(* Logix 5000 project; controller PLC_MCC1300_75F1 vendor 1 type 14 code 166 rev 32.11; software revision 32.04; part 17 of 83 *)
(* tags used below, declared in another part *)
   M302SpeedUp : MAC_SpeedUp;
   TMP_d : DINT;
   TMP_xPositioning : BOOL;
   TMP_xReverse : BOOL;
   TMP_xRun : BOOL;
   xAlwaysOFF : BOOL;
   Z300_Conveyor : UDT_StandConv[29];
   Z300_Conveyor_Conf : UDT_Conveyor_Config[29];
   Z300_Conveyor_HMW : MAC_Conveyor_ZC_HMW[29];
   Z300_Conveyor_IN_MOTION : MAC_Conveyor_ZC_IN_MOTION[29];
   Z301_HMR : MAC_Zone_ML_HMR;
(* CommandLogic, continued *)

ROUTINE M307BM1_Conveyor_Output   (* ladder *)
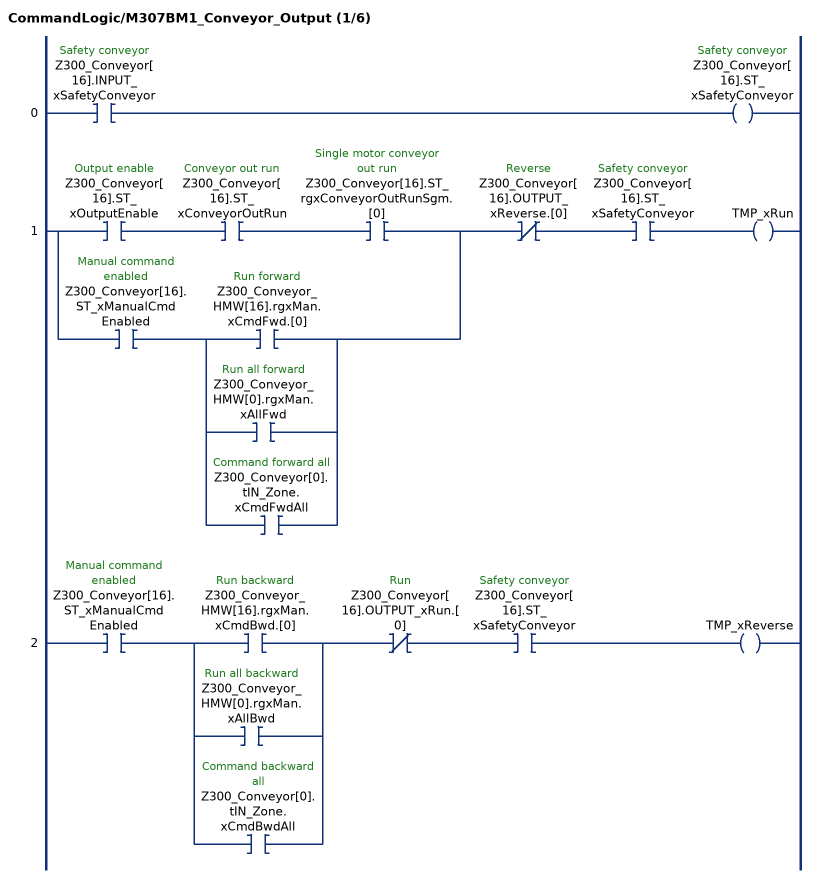
   0: XIC(Z300_Conveyor[16].INPUT_xSafetyConveyor)OTE(Z300_Conveyor[16].ST_xSafetyConveyor);
   1: [XIC(Z300_Conveyor[16].ST_xOutputEnable) XIC(Z300_Conveyor[16].ST_xConveyorOutRun) XIC(Z300_Conveyor[16].ST_rgxConveyorOutRunSgm.[0]) ,XIC(Z300_Conveyor[16].ST_xManualCmdEnabled) [XIC(Z300_Conveyor_HMW[16].rgxMan.xCmdFwd.[0]) ,XIC(Z300_Conveyor_HMW[0].rgxMan.xAllFwd) ,XIC(Z300_Conveyor[0].tIN_Zone.xCmdFwdAll) ] ]XIO(Z300_Conveyor[16].OUTPUT_xReverse.[0])XIC(Z300_Conveyor[16].ST_xSafetyConveyor)OTE(TMP_xRun);
   2: XIC(Z300_Conveyor[16].ST_xManualCmdEnabled)[XIC(Z300_Conveyor_HMW[16].rgxMan.xCmdBwd.[0]) ,XIC(Z300_Conveyor_HMW[0].rgxMan.xAllBwd) ,XIC(Z300_Conveyor[0].tIN_Zone.xCmdBwdAll) ]XIO(Z300_Conveyor[16].OUTPUT_xRun.[0])XIC(Z300_Conveyor[16].ST_xSafetyConveyor)OTE(TMP_xReverse);
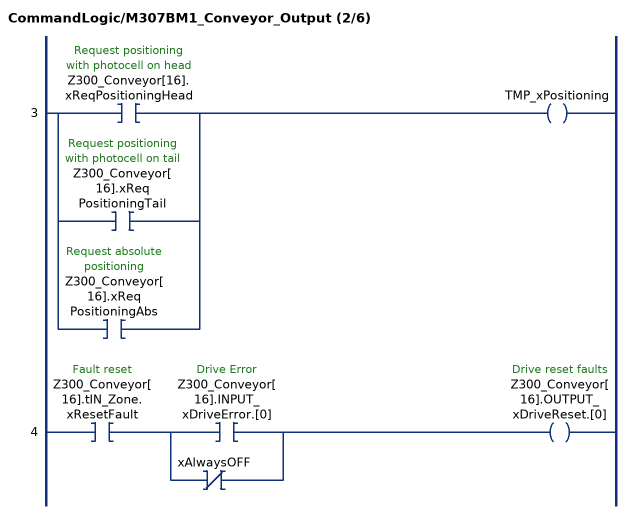
   3: [XIC(Z300_Conveyor[16].xReqPositioningHead) ,XIC(Z300_Conveyor[16].xReqPositioningTail) ,XIC(Z300_Conveyor[16].xReqPositioningAbs) ]OTE(TMP_xPositioning);
   4: XIC(Z300_Conveyor[16].tIN_Zone.xResetFault)[XIC(Z300_Conveyor[16].INPUT_xDriveError.[0]) ,XIO(xAlwaysOFF) ]OTE(Z300_Conveyor[16].OUTPUT_xDriveReset.[0]);
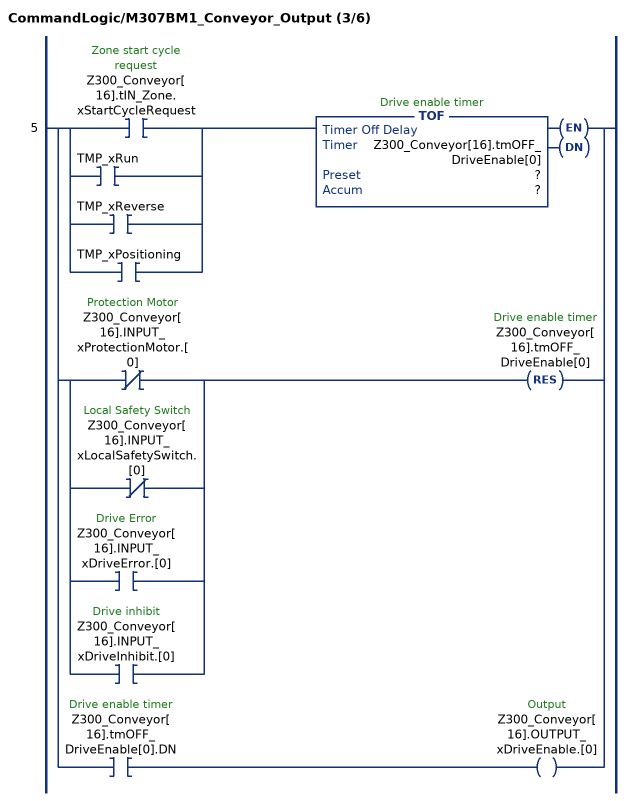
   5: [[XIC(Z300_Conveyor[16].tIN_Zone.xStartCycleRequest) ,XIC(TMP_xRun) ,XIC(TMP_xReverse) ,XIC(TMP_xPositioning) ] TOF(Z300_Conveyor[16].tmOFF_DriveEnable[0],?,?) ,[XIO(Z300_Conveyor[16].INPUT_xProtectionMotor.[0]) ,XIO(Z300_Conveyor[16].INPUT_xLocalSafetySwitch.[0]) ,XIC(Z300_Conveyor[16].INPUT_xDriveError.[0]) ,XIC(Z300_Conveyor[16].INPUT_xDriveInhibit.[0]) ] RES(Z300_Conveyor[16].tmOFF_DriveEnable[0]) ,XIC(Z300_Conveyor[16].tmOFF_DriveEnable[0].DN) OTE(Z300_Conveyor[16].OUTPUT_xDriveEnable.[0]) ];
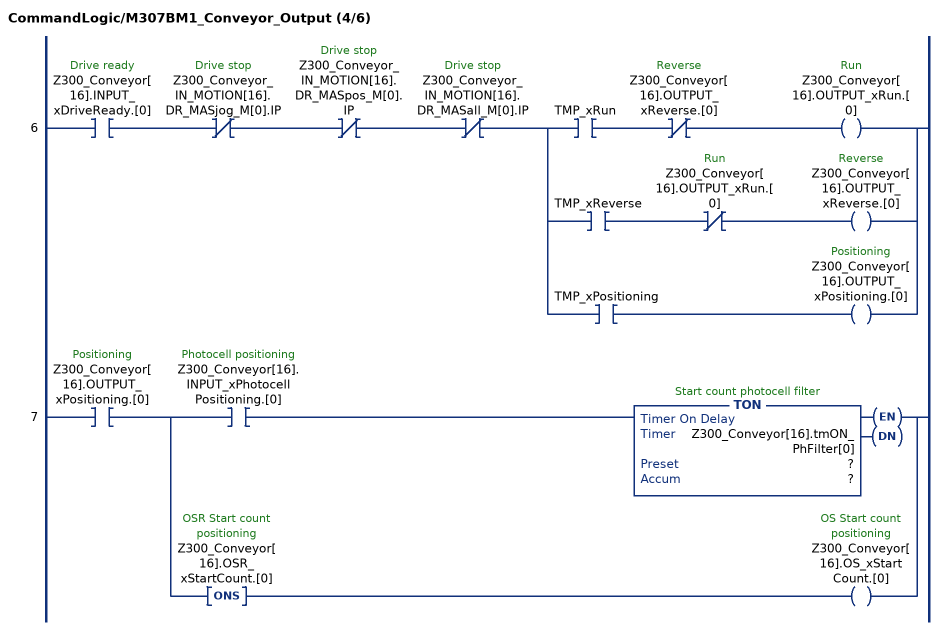
   6: XIC(Z300_Conveyor[16].INPUT_xDriveReady.[0])XIO(Z300_Conveyor_IN_MOTION[16].DR_MASjog_M[0].IP)XIO(Z300_Conveyor_IN_MOTION[16].DR_MASpos_M[0].IP)XIO(Z300_Conveyor_IN_MOTION[16].DR_MASall_M[0].IP)[XIC(TMP_xRun) XIO(Z300_Conveyor[16].OUTPUT_xReverse.[0]) OTE(Z300_Conveyor[16].OUTPUT_xRun.[0]) ,XIC(TMP_xReverse) XIO(Z300_Conveyor[16].OUTPUT_xRun.[0]) OTE(Z300_Conveyor[16].OUTPUT_xReverse.[0]) ,XIC(TMP_xPositioning) OTE(Z300_Conveyor[16].OUTPUT_xPositioning.[0]) ];
   7: XIC(Z300_Conveyor[16].OUTPUT_xPositioning.[0])[XIC(Z300_Conveyor[16].INPUT_xPhotocellPositioning.[0]) TON(Z300_Conveyor[16].tmON_PhFilter[0],?,?) ,ONS(Z300_Conveyor[16].OSR_xStartCount.[0]) OTE(Z300_Conveyor[16].OS_xStartCount.[0]) ];
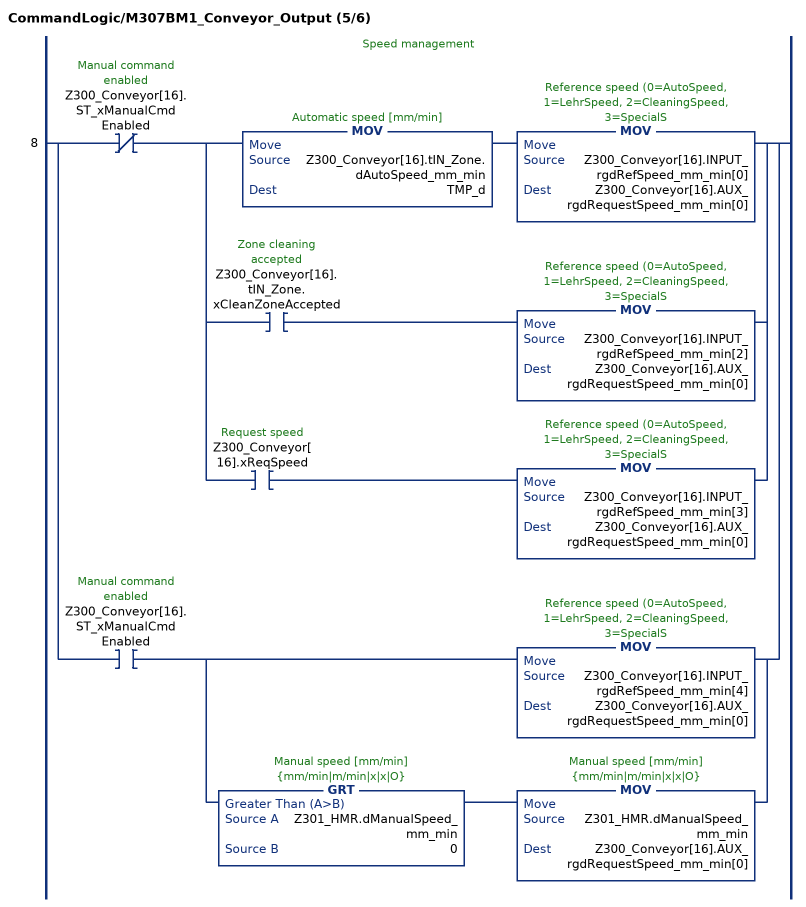
   // Speed management
   8: [XIO(Z300_Conveyor[16].ST_xManualCmdEnabled) [MOV(Z300_Conveyor[16].tIN_Zone.dAutoSpeed_mm_min,TMP_d) MOV(Z300_Conveyor[16].INPUT_rgdRefSpeed_mm_min[0],Z300_Conveyor[16].AUX_rgdRequestSpeed_mm_min[0]) ,XIC(Z300_Conveyor[16].tIN_Zone.xCleanZoneAccepted) MOV(Z300_Conveyor[16].INPUT_rgdRefSpeed_mm_min[2],Z300_Conveyor[16].AUX_rgdRequestSpeed_mm_min[0]) ,XIC(Z300_Conveyor[16].xReqSpeed) MOV(Z300_Conveyor[16].INPUT_rgdRefSpeed_mm_min[3],Z300_Conveyor[16].AUX_rgdRequestSpeed_mm_min[0]) ] ,XIC(Z300_Conveyor[16].ST_xManualCmdEnabled) [MOV(Z300_Conveyor[16].INPUT_rgdRefSpeed_mm_min[4],Z300_Conveyor[16].AUX_rgdRequestSpeed_mm_min[0]) ,GRT(Z301_HMR.dManualSpeed_mm_min,0) MOV(Z301_HMR.dManualSpeed_mm_min,Z300_Conveyor[16].AUX_rgdRequestSpeed_mm_min[0]) ] ];
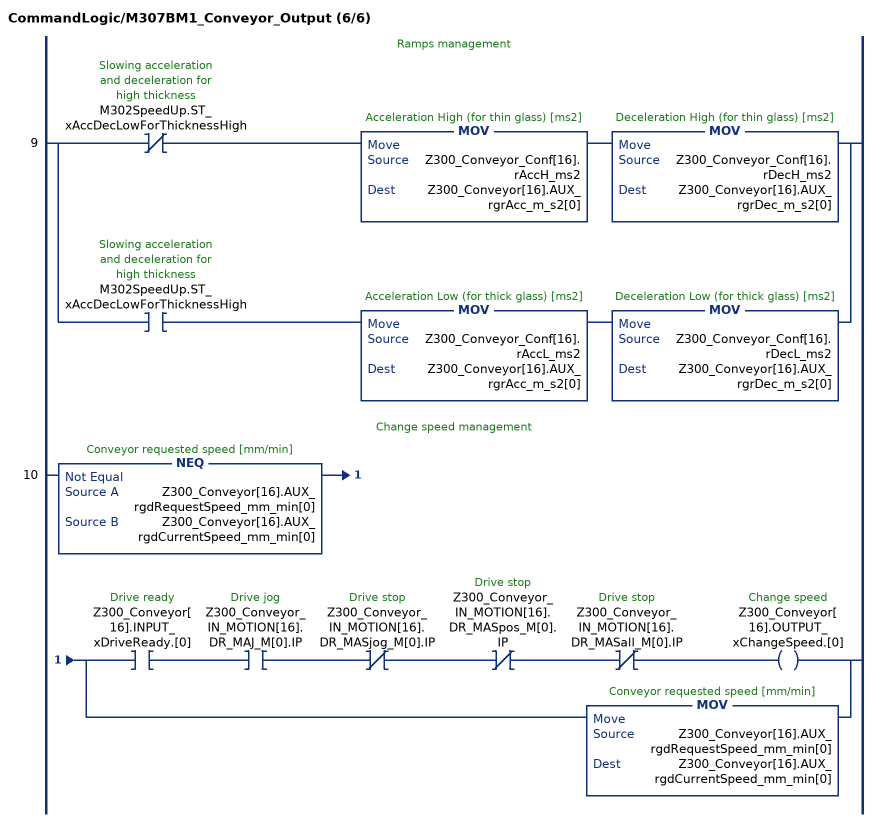
   // Ramps management
   9: [XIO(M302SpeedUp.ST_xAccDecLowForThicknessHigh) MOV(Z300_Conveyor_Conf[16].rAccH_ms2,Z300_Conveyor[16].AUX_rgrAcc_m_s2[0]) MOV(Z300_Conveyor_Conf[16].rDecH_ms2,Z300_Conveyor[16].AUX_rgrDec_m_s2[0]) ,XIC(M302SpeedUp.ST_xAccDecLowForThicknessHigh) MOV(Z300_Conveyor_Conf[16].rAccL_ms2,Z300_Conveyor[16].AUX_rgrAcc_m_s2[0]) MOV(Z300_Conveyor_Conf[16].rDecL_ms2,Z300_Conveyor[16].AUX_rgrDec_m_s2[0]) ];
   // Change speed management
   10: NEQ(Z300_Conveyor[16].AUX_rgdRequestSpeed_mm_min[0],Z300_Conveyor[16].AUX_rgdCurrentSpeed_mm_min[0])[XIC(Z300_Conveyor[16].INPUT_xDriveReady.[0]) XIC(Z300_Conveyor_IN_MOTION[16].DR_MAJ_M[0].IP) XIO(Z300_Conveyor_IN_MOTION[16].DR_MASjog_M[0].IP) XIO(Z300_Conveyor_IN_MOTION[16].DR_MASpos_M[0].IP) XIO(Z300_Conveyor_IN_MOTION[16].DR_MASall_M[0].IP) OTE(Z300_Conveyor[16].OUTPUT_xChangeSpeed.[0]) ,MOV(Z300_Conveyor[16].AUX_rgdRequestSpeed_mm_min[0],Z300_Conveyor[16].AUX_rgdCurrentSpeed_mm_min[0]) ];
END_ROUTINE

ROUTINE M307CM1_Conveyor_Output   (* ladder *)
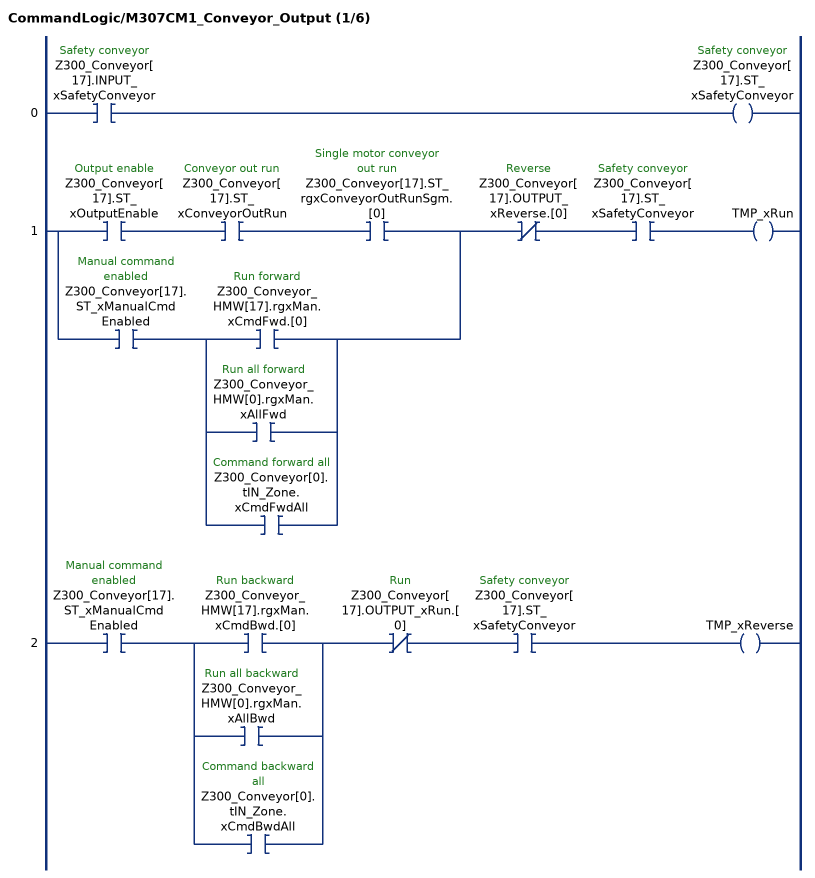
   0: XIC(Z300_Conveyor[17].INPUT_xSafetyConveyor)OTE(Z300_Conveyor[17].ST_xSafetyConveyor);
   1: [XIC(Z300_Conveyor[17].ST_xOutputEnable) XIC(Z300_Conveyor[17].ST_xConveyorOutRun) XIC(Z300_Conveyor[17].ST_rgxConveyorOutRunSgm.[0]) ,XIC(Z300_Conveyor[17].ST_xManualCmdEnabled) [XIC(Z300_Conveyor_HMW[17].rgxMan.xCmdFwd.[0]) ,XIC(Z300_Conveyor_HMW[0].rgxMan.xAllFwd) ,XIC(Z300_Conveyor[0].tIN_Zone.xCmdFwdAll) ] ]XIO(Z300_Conveyor[17].OUTPUT_xReverse.[0])XIC(Z300_Conveyor[17].ST_xSafetyConveyor)OTE(TMP_xRun);
   2: XIC(Z300_Conveyor[17].ST_xManualCmdEnabled)[XIC(Z300_Conveyor_HMW[17].rgxMan.xCmdBwd.[0]) ,XIC(Z300_Conveyor_HMW[0].rgxMan.xAllBwd) ,XIC(Z300_Conveyor[0].tIN_Zone.xCmdBwdAll) ]XIO(Z300_Conveyor[17].OUTPUT_xRun.[0])XIC(Z300_Conveyor[17].ST_xSafetyConveyor)OTE(TMP_xReverse);
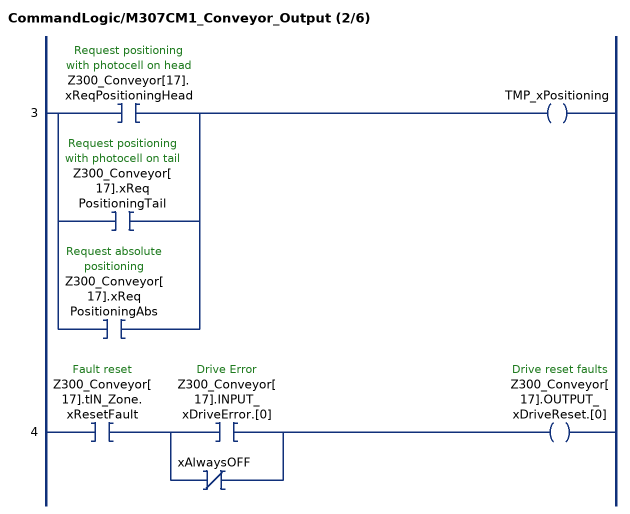
   3: [XIC(Z300_Conveyor[17].xReqPositioningHead) ,XIC(Z300_Conveyor[17].xReqPositioningTail) ,XIC(Z300_Conveyor[17].xReqPositioningAbs) ]OTE(TMP_xPositioning);
   4: XIC(Z300_Conveyor[17].tIN_Zone.xResetFault)[XIC(Z300_Conveyor[17].INPUT_xDriveError.[0]) ,XIO(xAlwaysOFF) ]OTE(Z300_Conveyor[17].OUTPUT_xDriveReset.[0]);
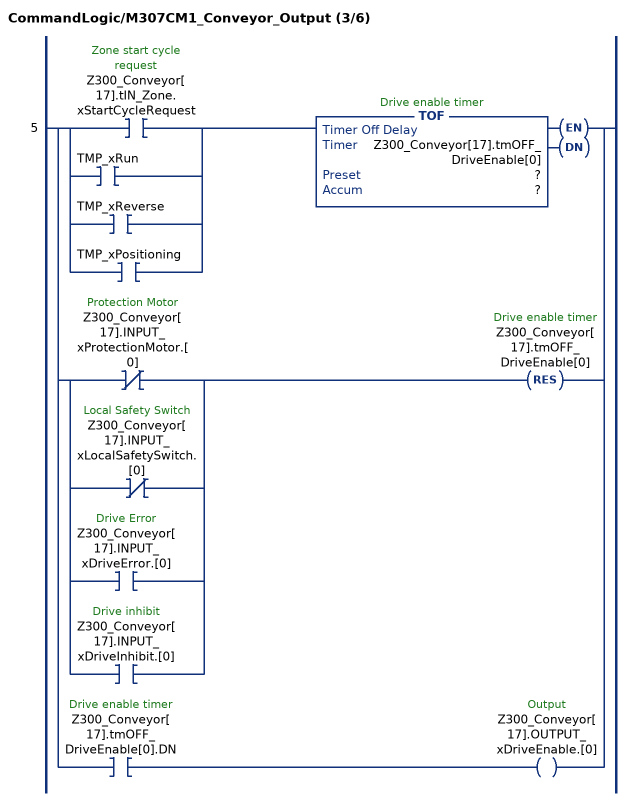
   5: [[XIC(Z300_Conveyor[17].tIN_Zone.xStartCycleRequest) ,XIC(TMP_xRun) ,XIC(TMP_xReverse) ,XIC(TMP_xPositioning) ] TOF(Z300_Conveyor[17].tmOFF_DriveEnable[0],?,?) ,[XIO(Z300_Conveyor[17].INPUT_xProtectionMotor.[0]) ,XIO(Z300_Conveyor[17].INPUT_xLocalSafetySwitch.[0]) ,XIC(Z300_Conveyor[17].INPUT_xDriveError.[0]) ,XIC(Z300_Conveyor[17].INPUT_xDriveInhibit.[0]) ] RES(Z300_Conveyor[17].tmOFF_DriveEnable[0]) ,XIC(Z300_Conveyor[17].tmOFF_DriveEnable[0].DN) OTE(Z300_Conveyor[17].OUTPUT_xDriveEnable.[0]) ];
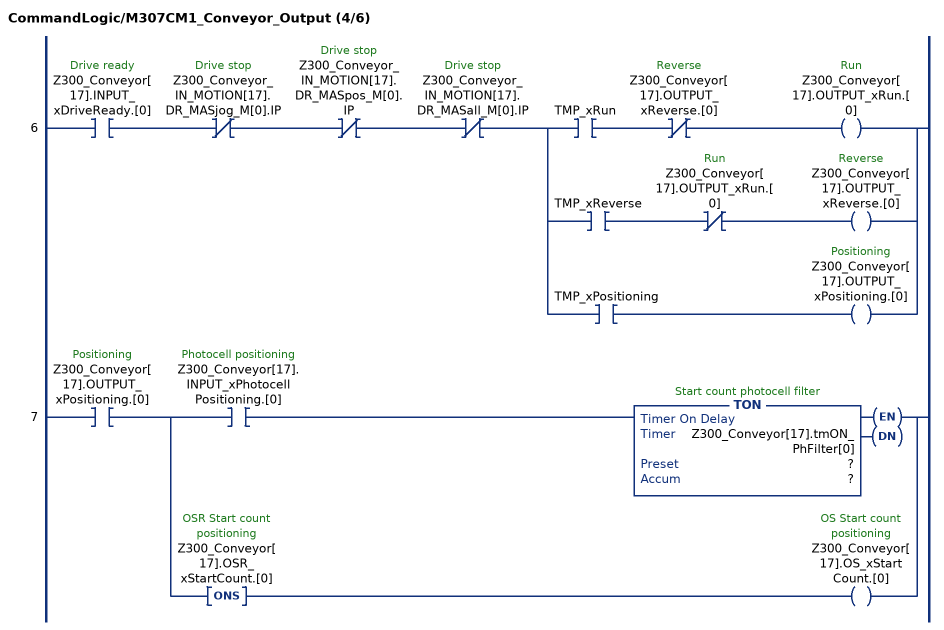
   6: XIC(Z300_Conveyor[17].INPUT_xDriveReady.[0])XIO(Z300_Conveyor_IN_MOTION[17].DR_MASjog_M[0].IP)XIO(Z300_Conveyor_IN_MOTION[17].DR_MASpos_M[0].IP)XIO(Z300_Conveyor_IN_MOTION[17].DR_MASall_M[0].IP)[XIC(TMP_xRun) XIO(Z300_Conveyor[17].OUTPUT_xReverse.[0]) OTE(Z300_Conveyor[17].OUTPUT_xRun.[0]) ,XIC(TMP_xReverse) XIO(Z300_Conveyor[17].OUTPUT_xRun.[0]) OTE(Z300_Conveyor[17].OUTPUT_xReverse.[0]) ,XIC(TMP_xPositioning) OTE(Z300_Conveyor[17].OUTPUT_xPositioning.[0]) ];
   7: XIC(Z300_Conveyor[17].OUTPUT_xPositioning.[0])[XIC(Z300_Conveyor[17].INPUT_xPhotocellPositioning.[0]) TON(Z300_Conveyor[17].tmON_PhFilter[0],?,?) ,ONS(Z300_Conveyor[17].OSR_xStartCount.[0]) OTE(Z300_Conveyor[17].OS_xStartCount.[0]) ];
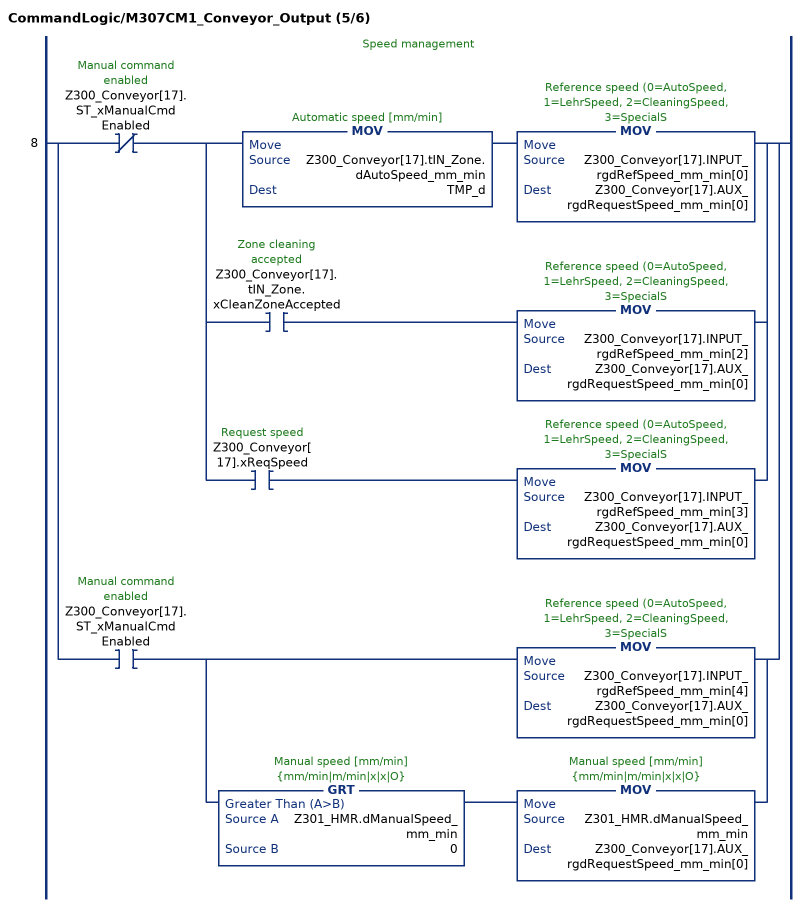
   // Speed management
   8: [XIO(Z300_Conveyor[17].ST_xManualCmdEnabled) [MOV(Z300_Conveyor[17].tIN_Zone.dAutoSpeed_mm_min,TMP_d) MOV(Z300_Conveyor[17].INPUT_rgdRefSpeed_mm_min[0],Z300_Conveyor[17].AUX_rgdRequestSpeed_mm_min[0]) ,XIC(Z300_Conveyor[17].tIN_Zone.xCleanZoneAccepted) MOV(Z300_Conveyor[17].INPUT_rgdRefSpeed_mm_min[2],Z300_Conveyor[17].AUX_rgdRequestSpeed_mm_min[0]) ,XIC(Z300_Conveyor[17].xReqSpeed) MOV(Z300_Conveyor[17].INPUT_rgdRefSpeed_mm_min[3],Z300_Conveyor[17].AUX_rgdRequestSpeed_mm_min[0]) ] ,XIC(Z300_Conveyor[17].ST_xManualCmdEnabled) [MOV(Z300_Conveyor[17].INPUT_rgdRefSpeed_mm_min[4],Z300_Conveyor[17].AUX_rgdRequestSpeed_mm_min[0]) ,GRT(Z301_HMR.dManualSpeed_mm_min,0) MOV(Z301_HMR.dManualSpeed_mm_min,Z300_Conveyor[17].AUX_rgdRequestSpeed_mm_min[0]) ] ];
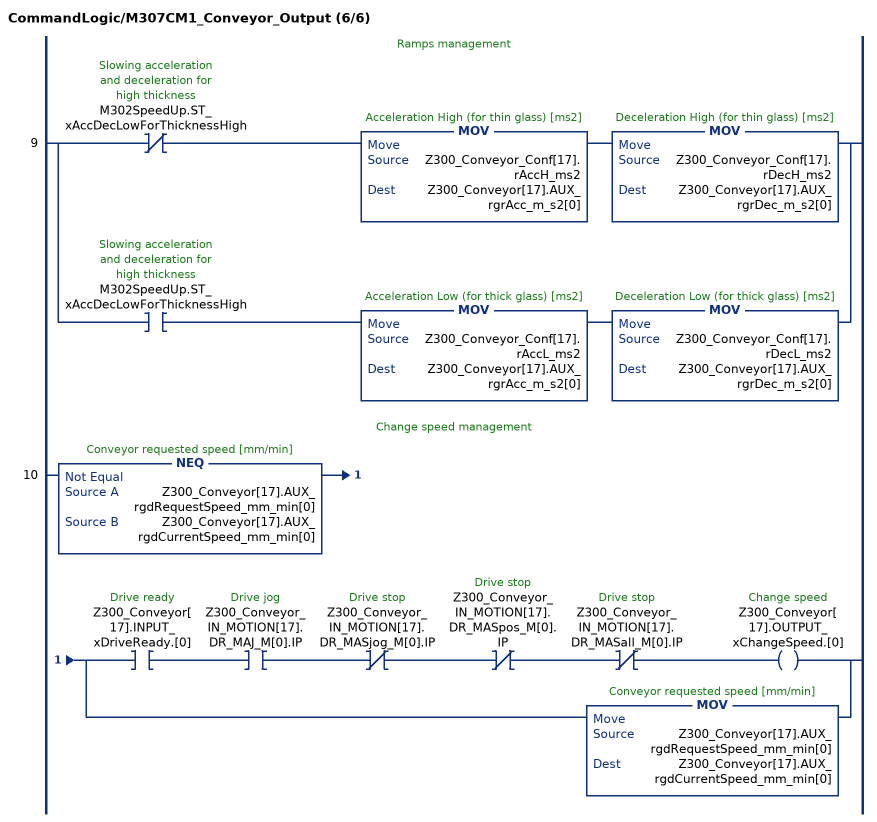
   // Ramps management
   9: [XIO(M302SpeedUp.ST_xAccDecLowForThicknessHigh) MOV(Z300_Conveyor_Conf[17].rAccH_ms2,Z300_Conveyor[17].AUX_rgrAcc_m_s2[0]) MOV(Z300_Conveyor_Conf[17].rDecH_ms2,Z300_Conveyor[17].AUX_rgrDec_m_s2[0]) ,XIC(M302SpeedUp.ST_xAccDecLowForThicknessHigh) MOV(Z300_Conveyor_Conf[17].rAccL_ms2,Z300_Conveyor[17].AUX_rgrAcc_m_s2[0]) MOV(Z300_Conveyor_Conf[17].rDecL_ms2,Z300_Conveyor[17].AUX_rgrDec_m_s2[0]) ];
   // Change speed management
   10: NEQ(Z300_Conveyor[17].AUX_rgdRequestSpeed_mm_min[0],Z300_Conveyor[17].AUX_rgdCurrentSpeed_mm_min[0])[XIC(Z300_Conveyor[17].INPUT_xDriveReady.[0]) XIC(Z300_Conveyor_IN_MOTION[17].DR_MAJ_M[0].IP) XIO(Z300_Conveyor_IN_MOTION[17].DR_MASjog_M[0].IP) XIO(Z300_Conveyor_IN_MOTION[17].DR_MASpos_M[0].IP) XIO(Z300_Conveyor_IN_MOTION[17].DR_MASall_M[0].IP) OTE(Z300_Conveyor[17].OUTPUT_xChangeSpeed.[0]) ,MOV(Z300_Conveyor[17].AUX_rgdRequestSpeed_mm_min[0],Z300_Conveyor[17].AUX_rgdCurrentSpeed_mm_min[0]) ];
END_ROUTINE

ROUTINE M307DM1_Conveyor_Output   (* ladder *)
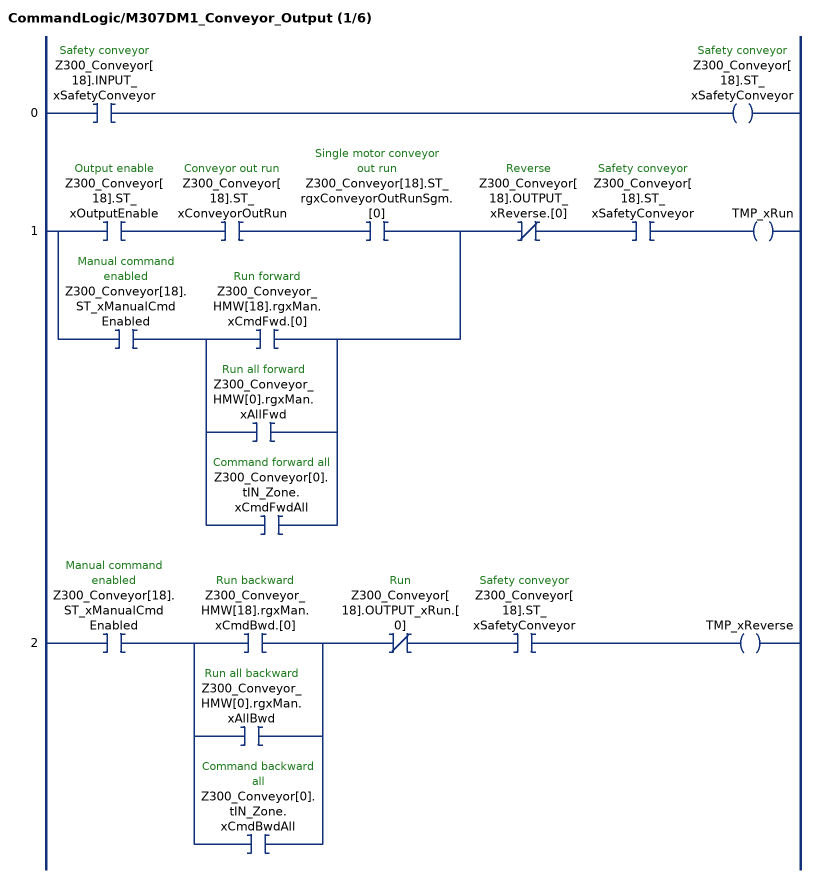
   0: XIC(Z300_Conveyor[18].INPUT_xSafetyConveyor)OTE(Z300_Conveyor[18].ST_xSafetyConveyor);
   1: [XIC(Z300_Conveyor[18].ST_xOutputEnable) XIC(Z300_Conveyor[18].ST_xConveyorOutRun) XIC(Z300_Conveyor[18].ST_rgxConveyorOutRunSgm.[0]) ,XIC(Z300_Conveyor[18].ST_xManualCmdEnabled) [XIC(Z300_Conveyor_HMW[18].rgxMan.xCmdFwd.[0]) ,XIC(Z300_Conveyor_HMW[0].rgxMan.xAllFwd) ,XIC(Z300_Conveyor[0].tIN_Zone.xCmdFwdAll) ] ]XIO(Z300_Conveyor[18].OUTPUT_xReverse.[0])XIC(Z300_Conveyor[18].ST_xSafetyConveyor)OTE(TMP_xRun);
   2: XIC(Z300_Conveyor[18].ST_xManualCmdEnabled)[XIC(Z300_Conveyor_HMW[18].rgxMan.xCmdBwd.[0]) ,XIC(Z300_Conveyor_HMW[0].rgxMan.xAllBwd) ,XIC(Z300_Conveyor[0].tIN_Zone.xCmdBwdAll) ]XIO(Z300_Conveyor[18].OUTPUT_xRun.[0])XIC(Z300_Conveyor[18].ST_xSafetyConveyor)OTE(TMP_xReverse);
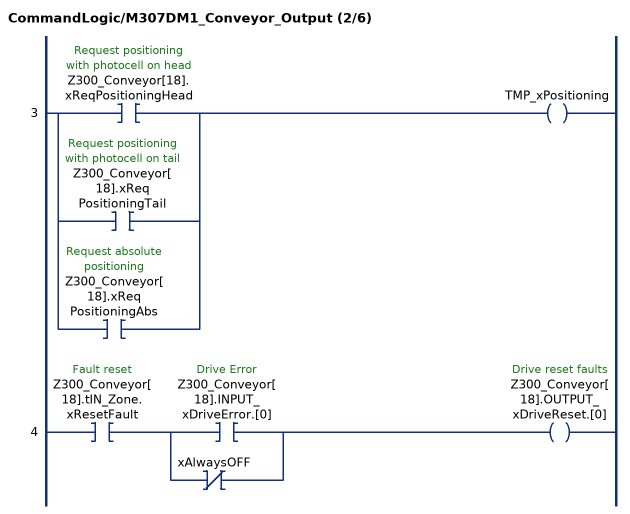
   3: [XIC(Z300_Conveyor[18].xReqPositioningHead) ,XIC(Z300_Conveyor[18].xReqPositioningTail) ,XIC(Z300_Conveyor[18].xReqPositioningAbs) ]OTE(TMP_xPositioning);
   4: XIC(Z300_Conveyor[18].tIN_Zone.xResetFault)[XIC(Z300_Conveyor[18].INPUT_xDriveError.[0]) ,XIO(xAlwaysOFF) ]OTE(Z300_Conveyor[18].OUTPUT_xDriveReset.[0]);
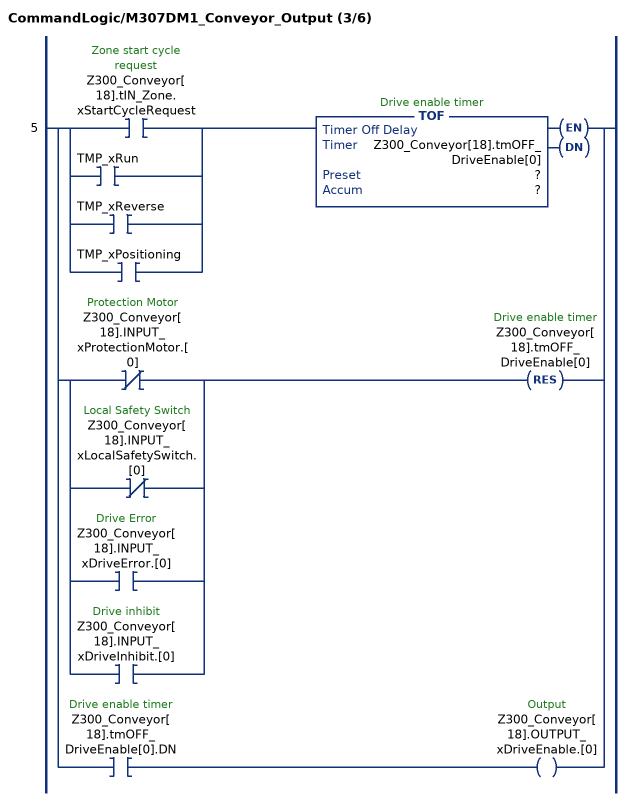
   5: [[XIC(Z300_Conveyor[18].tIN_Zone.xStartCycleRequest) ,XIC(TMP_xRun) ,XIC(TMP_xReverse) ,XIC(TMP_xPositioning) ] TOF(Z300_Conveyor[18].tmOFF_DriveEnable[0],?,?) ,[XIO(Z300_Conveyor[18].INPUT_xProtectionMotor.[0]) ,XIO(Z300_Conveyor[18].INPUT_xLocalSafetySwitch.[0]) ,XIC(Z300_Conveyor[18].INPUT_xDriveError.[0]) ,XIC(Z300_Conveyor[18].INPUT_xDriveInhibit.[0]) ] RES(Z300_Conveyor[18].tmOFF_DriveEnable[0]) ,XIC(Z300_Conveyor[18].tmOFF_DriveEnable[0].DN) OTE(Z300_Conveyor[18].OUTPUT_xDriveEnable.[0]) ];
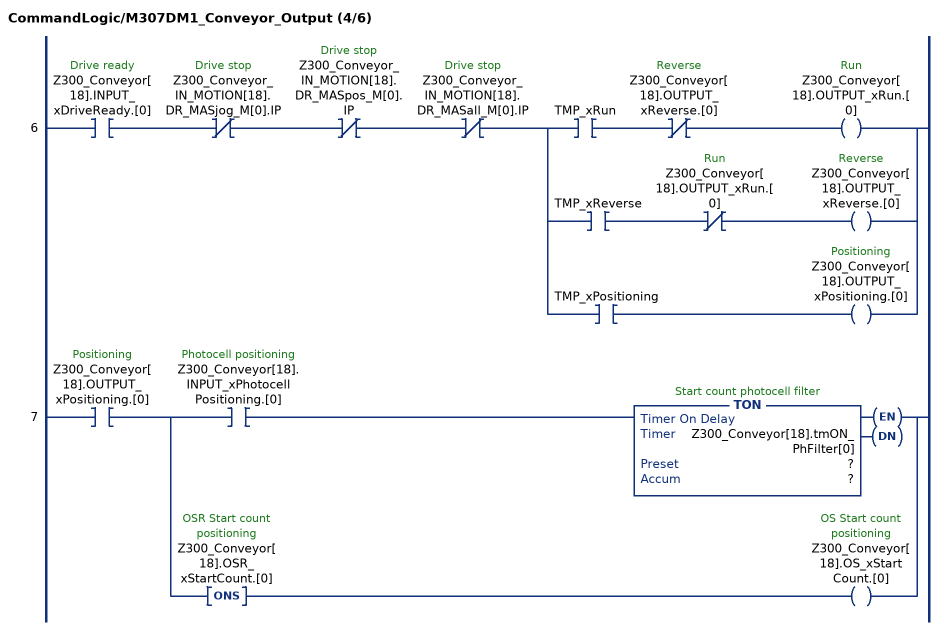
   6: XIC(Z300_Conveyor[18].INPUT_xDriveReady.[0])XIO(Z300_Conveyor_IN_MOTION[18].DR_MASjog_M[0].IP)XIO(Z300_Conveyor_IN_MOTION[18].DR_MASpos_M[0].IP)XIO(Z300_Conveyor_IN_MOTION[18].DR_MASall_M[0].IP)[XIC(TMP_xRun) XIO(Z300_Conveyor[18].OUTPUT_xReverse.[0]) OTE(Z300_Conveyor[18].OUTPUT_xRun.[0]) ,XIC(TMP_xReverse) XIO(Z300_Conveyor[18].OUTPUT_xRun.[0]) OTE(Z300_Conveyor[18].OUTPUT_xReverse.[0]) ,XIC(TMP_xPositioning) OTE(Z300_Conveyor[18].OUTPUT_xPositioning.[0]) ];
   7: XIC(Z300_Conveyor[18].OUTPUT_xPositioning.[0])[XIC(Z300_Conveyor[18].INPUT_xPhotocellPositioning.[0]) TON(Z300_Conveyor[18].tmON_PhFilter[0],?,?) ,ONS(Z300_Conveyor[18].OSR_xStartCount.[0]) OTE(Z300_Conveyor[18].OS_xStartCount.[0]) ];
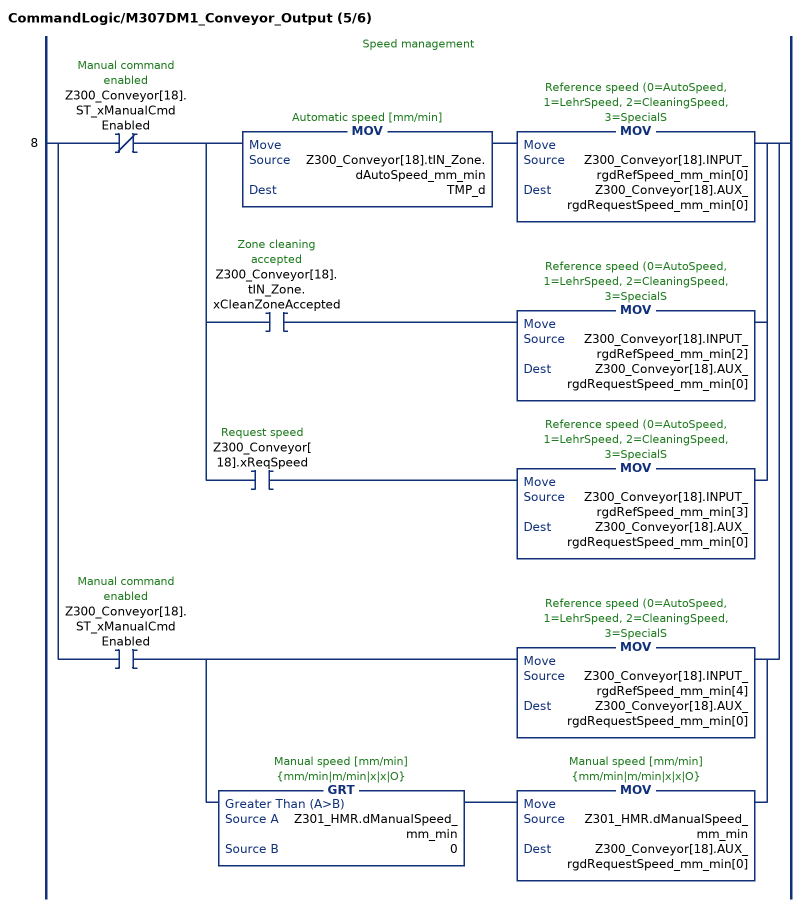
   // Speed management
   8: [XIO(Z300_Conveyor[18].ST_xManualCmdEnabled) [MOV(Z300_Conveyor[18].tIN_Zone.dAutoSpeed_mm_min,TMP_d) MOV(Z300_Conveyor[18].INPUT_rgdRefSpeed_mm_min[0],Z300_Conveyor[18].AUX_rgdRequestSpeed_mm_min[0]) ,XIC(Z300_Conveyor[18].tIN_Zone.xCleanZoneAccepted) MOV(Z300_Conveyor[18].INPUT_rgdRefSpeed_mm_min[2],Z300_Conveyor[18].AUX_rgdRequestSpeed_mm_min[0]) ,XIC(Z300_Conveyor[18].xReqSpeed) MOV(Z300_Conveyor[18].INPUT_rgdRefSpeed_mm_min[3],Z300_Conveyor[18].AUX_rgdRequestSpeed_mm_min[0]) ] ,XIC(Z300_Conveyor[18].ST_xManualCmdEnabled) [MOV(Z300_Conveyor[18].INPUT_rgdRefSpeed_mm_min[4],Z300_Conveyor[18].AUX_rgdRequestSpeed_mm_min[0]) ,GRT(Z301_HMR.dManualSpeed_mm_min,0) MOV(Z301_HMR.dManualSpeed_mm_min,Z300_Conveyor[18].AUX_rgdRequestSpeed_mm_min[0]) ] ];
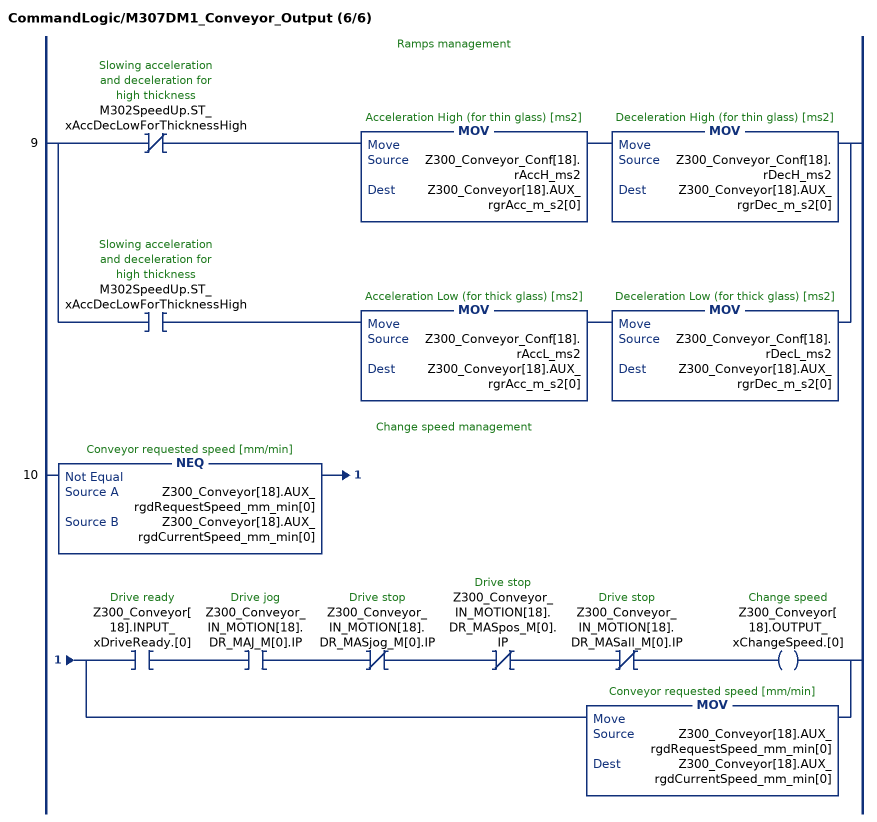
   // Ramps management
   9: [XIO(M302SpeedUp.ST_xAccDecLowForThicknessHigh) MOV(Z300_Conveyor_Conf[18].rAccH_ms2,Z300_Conveyor[18].AUX_rgrAcc_m_s2[0]) MOV(Z300_Conveyor_Conf[18].rDecH_ms2,Z300_Conveyor[18].AUX_rgrDec_m_s2[0]) ,XIC(M302SpeedUp.ST_xAccDecLowForThicknessHigh) MOV(Z300_Conveyor_Conf[18].rAccL_ms2,Z300_Conveyor[18].AUX_rgrAcc_m_s2[0]) MOV(Z300_Conveyor_Conf[18].rDecL_ms2,Z300_Conveyor[18].AUX_rgrDec_m_s2[0]) ];
   // Change speed management
   10: NEQ(Z300_Conveyor[18].AUX_rgdRequestSpeed_mm_min[0],Z300_Conveyor[18].AUX_rgdCurrentSpeed_mm_min[0])[XIC(Z300_Conveyor[18].INPUT_xDriveReady.[0]) XIC(Z300_Conveyor_IN_MOTION[18].DR_MAJ_M[0].IP) XIO(Z300_Conveyor_IN_MOTION[18].DR_MASjog_M[0].IP) XIO(Z300_Conveyor_IN_MOTION[18].DR_MASpos_M[0].IP) XIO(Z300_Conveyor_IN_MOTION[18].DR_MASall_M[0].IP) OTE(Z300_Conveyor[18].OUTPUT_xChangeSpeed.[0]) ,MOV(Z300_Conveyor[18].AUX_rgdRequestSpeed_mm_min[0],Z300_Conveyor[18].AUX_rgdCurrentSpeed_mm_min[0]) ];
END_ROUTINE
